// TIA Portal project "Lagerregal_3" (V20) (continued)
VERSION : 0.1
   VAR_INPUT
      eAutomatik : Bool;   // Automatikmodus
      eAusschalten : Bool;   // Ausschalten der Schrittkette
      T_1_2 : Bool;
      T_2_3 : Bool;
      T_3_4 : Bool := TRUE;
      T_4_5 : Bool := TRUE;
      T_5_6 : Bool := TRUE;
      T_6_7 : Bool := TRUE;
      T_7_8 : Bool := TRUE;
      T_8_9 : Bool := TRUE;
      T_9_10 : Bool := TRUE;
      T_10_1 : Bool := TRUE;
   END_VAR
   VAR_OUTPUT
      aSchrittnummer : Int;
   END_VAR
   VAR
      Step_1 : Bool;
      Step_2 : Bool;
      Step_3 : Bool;
      Step_4 : Bool;
      Step_5 : Bool;
      Step_6 : Bool;
      Step_7 : Bool;
      Step_8 : Bool;
      Step_9 : Bool;
      Step_10 : Bool;
   END_VAR
BEGIN

REGION Network 1: Step 1
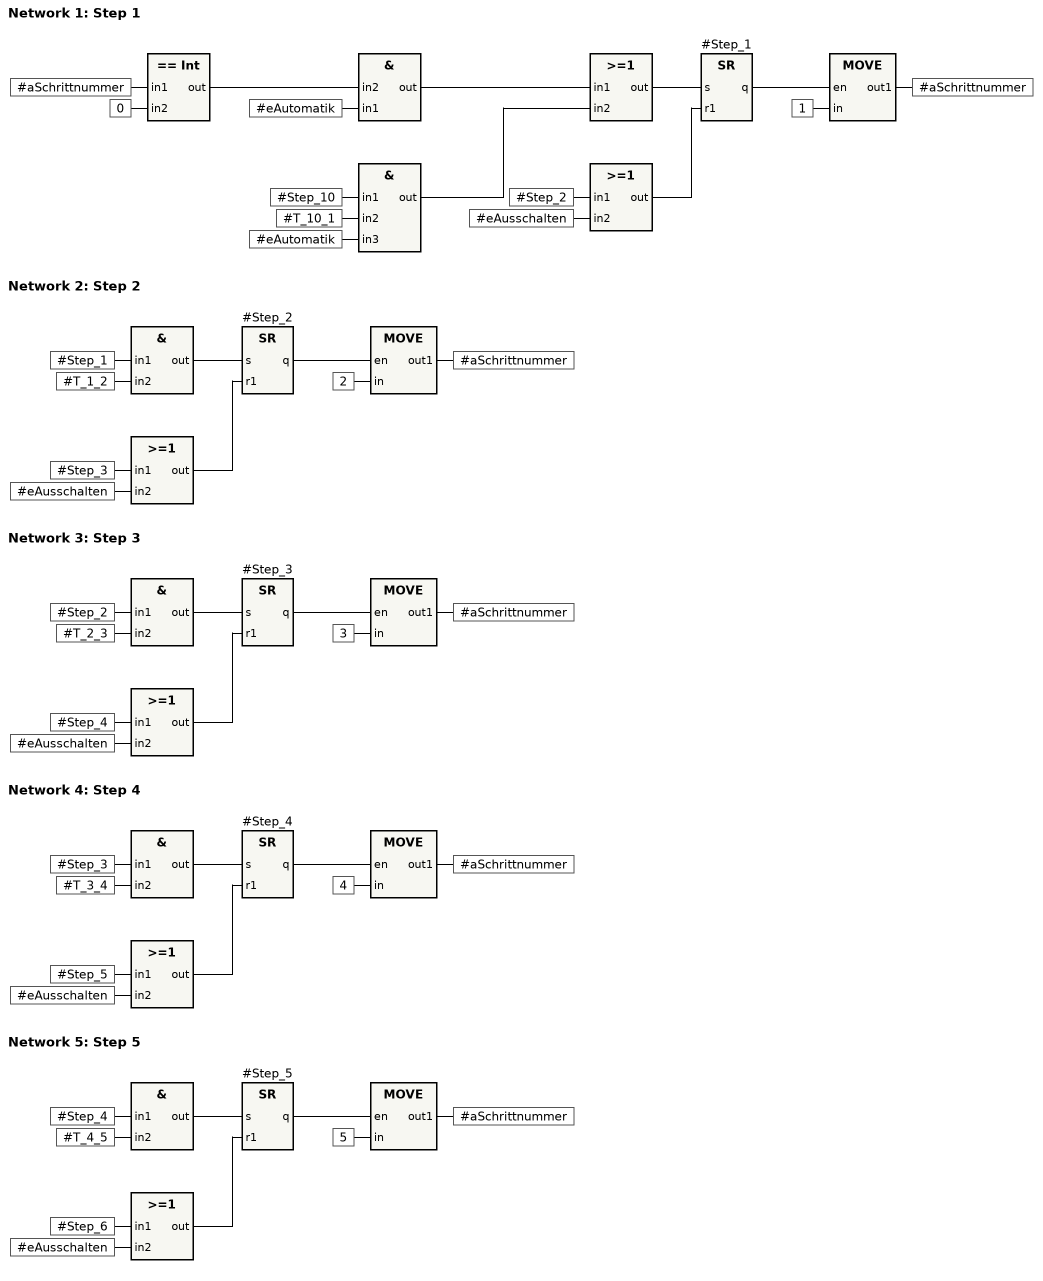
   IF ((#aSchrittnummer = 0) AND #eAutomatik) OR (#Step_10 AND #T_10_1 AND #eAutomatik) THEN
       #Step_1 := TRUE;   // SR flip-flop
   END_IF;
   IF #Step_2 OR #eAusschalten THEN #Step_1 := FALSE; END_IF;
   IF #Step_1 THEN #aSchrittnummer := 1; END_IF;
END_REGION

REGION Network 2: Step 2
   IF #Step_1 AND #T_1_2 THEN
       #Step_2 := TRUE;   // SR flip-flop
   END_IF;
   IF #Step_3 OR #eAusschalten THEN #Step_2 := FALSE; END_IF;
   IF #Step_2 THEN #aSchrittnummer := 2; END_IF;
END_REGION

REGION Network 3: Step 3
   IF #Step_2 AND #T_2_3 THEN
       #Step_3 := TRUE;   // SR flip-flop
   END_IF;
   IF #Step_4 OR #eAusschalten THEN #Step_3 := FALSE; END_IF;
   IF #Step_3 THEN #aSchrittnummer := 3; END_IF;
END_REGION

REGION Network 4: Step 4
   IF #Step_3 AND #T_3_4 THEN
       #Step_4 := TRUE;   // SR flip-flop
   END_IF;
   IF #Step_5 OR #eAusschalten THEN #Step_4 := FALSE; END_IF;
   IF #Step_4 THEN #aSchrittnummer := 4; END_IF;
END_REGION

REGION Network 5: Step 5
   IF #Step_4 AND #T_4_5 THEN
       #Step_5 := TRUE;   // SR flip-flop
   END_IF;
   IF #Step_6 OR #eAusschalten THEN #Step_5 := FALSE; END_IF;
   IF #Step_5 THEN #aSchrittnummer := 5; END_IF;
END_REGION

REGION Network 6: Step 6
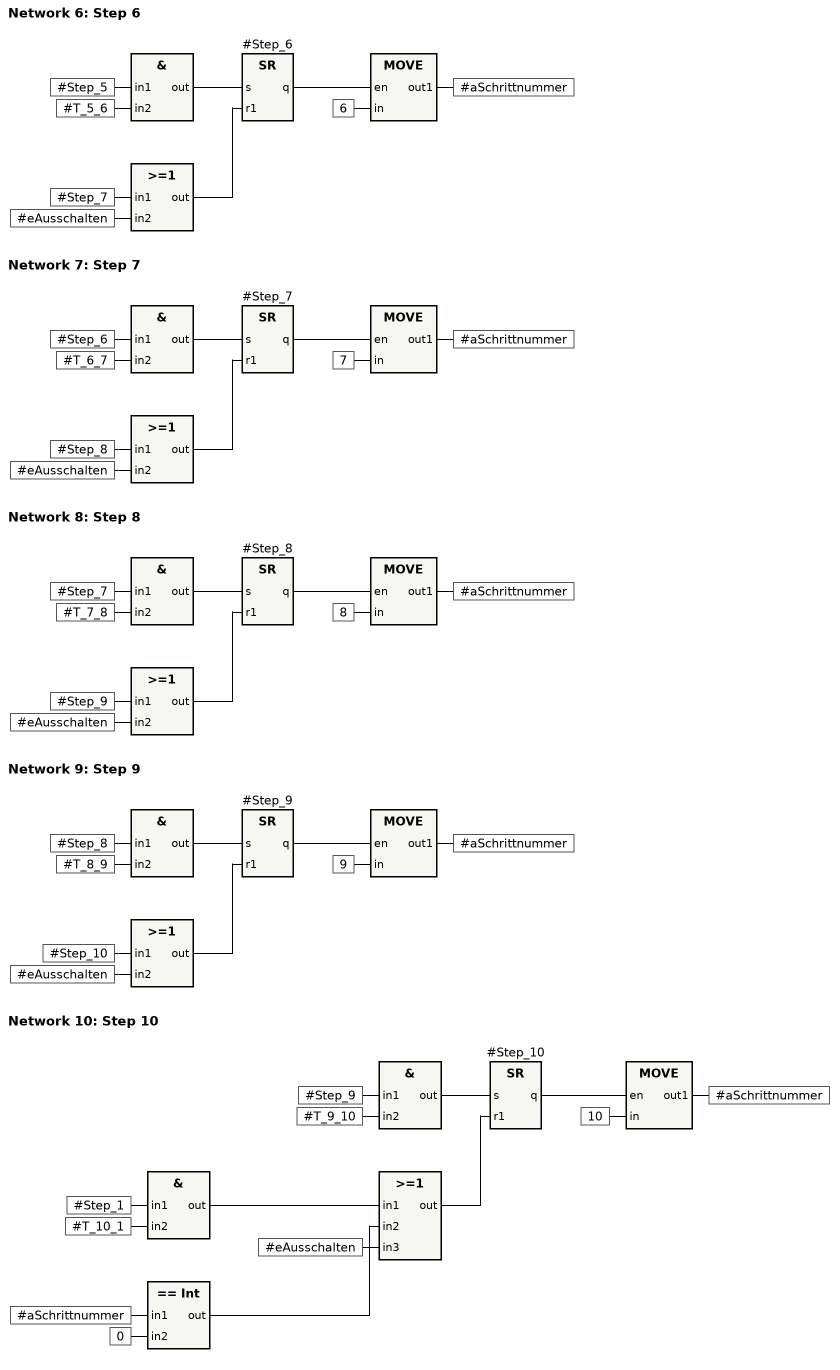
   IF #Step_5 AND #T_5_6 THEN
       #Step_6 := TRUE;   // SR flip-flop
   END_IF;
   IF #Step_7 OR #eAusschalten THEN #Step_6 := FALSE; END_IF;
   IF #Step_6 THEN #aSchrittnummer := 6; END_IF;
END_REGION

REGION Network 7: Step 7
   IF #Step_6 AND #T_6_7 THEN
       #Step_7 := TRUE;   // SR flip-flop
   END_IF;
   IF #Step_8 OR #eAusschalten THEN #Step_7 := FALSE; END_IF;
   IF #Step_7 THEN #aSchrittnummer := 7; END_IF;
END_REGION

REGION Network 8: Step 8
   IF #Step_7 AND #T_7_8 THEN
       #Step_8 := TRUE;   // SR flip-flop
   END_IF;
   IF #Step_9 OR #eAusschalten THEN #Step_8 := FALSE; END_IF;
   IF #Step_8 THEN #aSchrittnummer := 8; END_IF;
END_REGION

REGION Network 9: Step 9
   IF #Step_8 AND #T_8_9 THEN
       #Step_9 := TRUE;   // SR flip-flop
   END_IF;
   IF #Step_10 OR #eAusschalten THEN #Step_9 := FALSE; END_IF;
   IF #Step_9 THEN #aSchrittnummer := 9; END_IF;
END_REGION

REGION Network 10: Step 10
   IF #Step_9 AND #T_9_10 THEN
       #Step_10 := TRUE;   // SR flip-flop
   END_IF;
   IF (#Step_1 AND #T_10_1) OR (#aSchrittnummer = 0) OR #eAusschalten THEN #Step_10 := FALSE; END_IF;
   IF #Step_10 THEN #aSchrittnummer := 10; END_IF;
END_REGION

REGION Network 11: Schrittkette beenden, wenn der Automatikmodus beendet wird
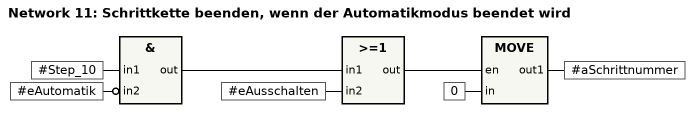
   IF (#Step_10 AND NOT #eAutomatik) OR #eAusschalten THEN #aSchrittnummer := 0; END_IF;
END_REGION
END_FUNCTION_BLOCK

FUNCTION "Aus_Anlage" : Void   // FC1, FBD
{ S7_Optimized_Access := 'TRUE' }
VERSION : 0.1
BEGIN

REGION Network 1 (SCL): Gabelsteuerung Kran_1
   "6M1" := "HMI_Schnittstelle".Ausgaenge."6M1";
   "6M2" := "HMI_Schnittstelle".Ausgaenge."6M2";
END_REGION

REGION Network 2 (SCL): Gabelsteuerung Kran_2
   "7M1" := "HMI_Schnittstelle".Ausgaenge."7M1";
   "7M2" := "HMI_Schnittstelle".Ausgaenge."7M2";
END_REGION

REGION Network 3 (SCL): Foerderbaender Einlass
   "1M1" := "HMI_Schnittstelle".Ausgaenge."1M1";
   "2M1" := "HMI_Schnittstelle".Ausgaenge."2M1";
   "3M1" := "HMI_Schnittstelle".Ausgaenge."3M1";
END_REGION

REGION Network 4 (SCL): Foerderbaender Auslass
   "4M1" := "HMI_Schnittstelle".Ausgaenge."4M1";
   "5M1" := "HMI_Schnittstelle".Ausgaenge."5M1";
END_REGION

REGION Network 5 (SCL): Leuchte Starttaster
   "HMI_Schnittstelle".Ausgaenge.H1 := "HMI_Schnittstelle".Eingaenge.S2;
END_REGION
END_FUNCTION

FUNCTION "Aus_HMI" : Void   // FC20, FBD
{ S7_Optimized_Access := 'TRUE' }
VERSION : 0.1
BEGIN
END_FUNCTION

FUNCTION "Aus_Kran" : Void   // FC30, SCL
{ S7_Optimized_Access := 'TRUE' }
VERSION : 0.1
   VAR_INPUT
      "eX-Soll" : Int;
      "eZ-Soll" : Int;
      eGabel_links : Bool;
      eGabel_rechts : Bool;
   END_VAR
   VAR_OUTPUT
      aKran_X : Int;
      aKran_Z : Int;
      aKran_Gabel_links : Bool;
      aKran_Gabel_rechts : Bool;
   END_VAR
BEGIN
   // Kran Gabel
   #aKran_Gabel_links := #eGabel_links;
   #aKran_Gabel_rechts := #eGabel_rechts;


   // Kran Position
   // Kran X-Soll-Position
   #"aKran_X" := #"eX-Soll";
   // Kran Z-Soll-Position
   #"aKran_Z" := #"eZ-Soll";
END_FUNCTION

FUNCTION "Ausgabe_Stapler_EIN" : Void   // FC70, FBD
{ S7_Optimized_Access := 'TRUE' }
VERSION : 0.1
BEGIN

REGION Network 1: Sollposition X
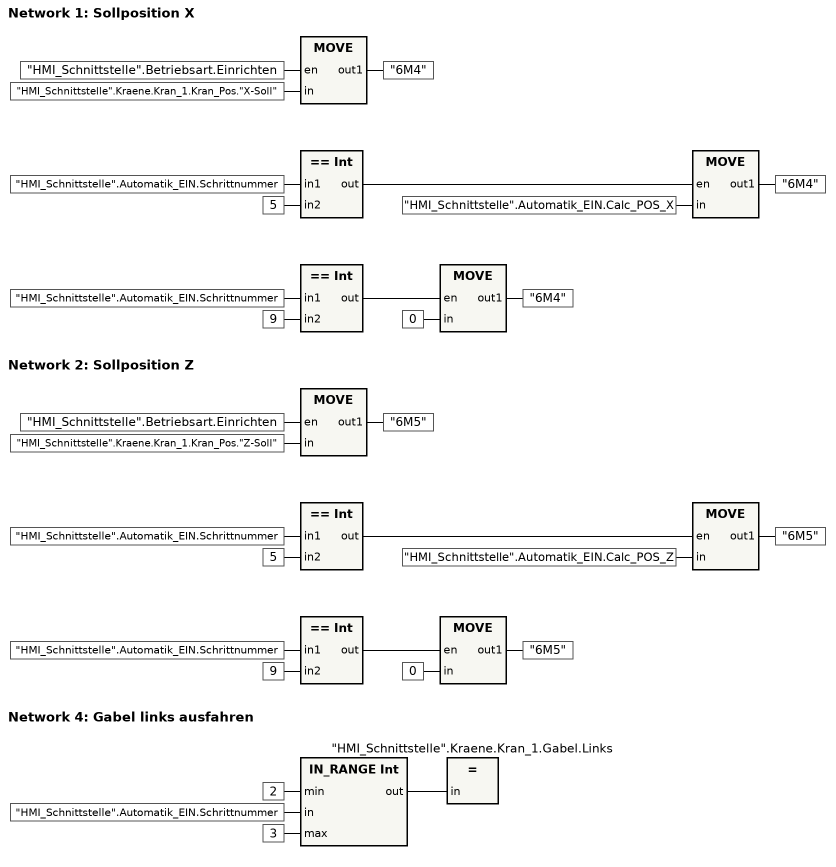
   IF "HMI_Schnittstelle".Betriebsart.Einrichten THEN
       "6M4" := "HMI_Schnittstelle".Kraene.Kran_1.Kran_Pos."X-Soll";
   END_IF;
   IF "HMI_Schnittstelle".Automatik_EIN.Schrittnummer = 5 THEN
       "6M4" := "HMI_Schnittstelle".Automatik_EIN.Calc_POS_X;
   END_IF;
   IF "HMI_Schnittstelle".Automatik_EIN.Schrittnummer = 9 THEN "6M4" := 0; END_IF;
END_REGION

REGION Network 2: Sollposition Z
   IF "HMI_Schnittstelle".Betriebsart.Einrichten THEN
       "6M5" := "HMI_Schnittstelle".Kraene.Kran_1.Kran_Pos."Z-Soll";
   END_IF;
   IF "HMI_Schnittstelle".Automatik_EIN.Schrittnummer = 5 THEN
       "6M5" := "HMI_Schnittstelle".Automatik_EIN.Calc_POS_Z;
   END_IF;
   IF "HMI_Schnittstelle".Automatik_EIN.Schrittnummer = 9 THEN "6M5" := 0; END_IF;
END_REGION

REGION Network 3 (SCL): Z-Achse Kran 1 Soll-Pos
   // Einrichtbetrieb
   IF "HMI_Schnittstelle".Betriebsart.Einrichten THEN
       "6M5" := "HMI_Schnittstelle".Kraene.Kran_1.Kran_Pos."Z-Soll";

   // Automatikbetrieb    
   ELSIF "HMI_Schnittstelle".Automatik_EIN.Schrittnummer = 3 THEN
       // Palette aus Grundstellung anheben
       "6M5" := "Anheben_Absenken" + 2;
   ELSIF "HMI_Schnittstelle".Automatik_EIN.Schrittnummer = 5 THEN
       //Fach mit Nummer anfahren
       "6M5" := "HMI_Schnittstelle".Automatik_EIN.Calc_POS_Z;
   ELSIF "HMI_Schnittstelle".Automatik_EIN.Schrittnummer = 7 THEN
       // Palette in Regal einlagern
       "6M5" := "HMI_Schnittstelle".Automatik_EIN.Calc_POS_Z - "Anheben_Absenken";
   ELSIF "HMI_Schnittstelle".Automatik_EIN.Schrittnummer = 9 THEN
       // Stapler in Grundstellung
       "6M5" := 0;
   END_IF;
END_REGION

REGION Network 4: Gabel links ausfahren
   "HMI_Schnittstelle".Kraene.Kran_1.Gabel.Links := (2 <= "HMI_Schnittstelle".Automatik_EIN.Schrittnummer) AND ("HMI_Schnittstelle".Automatik_EIN.Schrittnummer <= 3);
END_REGION

REGION Network 5 (SCL): Gabel rechts ausfahren
   "HMI_Schnittstelle".Kraene.Kran_1.Gabel.Rechts := "HMI_Schnittstelle".Automatik_EIN.Schrittnummer = 6
                                                   OR "HMI_Schnittstelle".Automatik_EIN.Schrittnummer = 7;
END_REGION
END_FUNCTION

FUNCTION "Berechne_Offset" : Void   // FC5000, SCL
{ S7_Optimized_Access := 'TRUE' }
VERSION : 0.1
   VAR_INPUT
      eFach_Nr : DInt;
      eFach_Anzahl : DInt;
      eFach_Breite : DInt;
      eFach_Hoehe : DInt;
      eOffset_X : DInt;
      eOffset_Z : DInt;
   END_VAR
   VAR_OUTPUT
      aPos_X : DInt;
      aPos_Z : DInt;
   END_VAR
BEGIN
   (*
      Der Baustein berechnet die Koordinaten (X,Z) eines Fachs
      in Abhängigkeit von einer Fachnummer

      Der Baustein ist universell einsetzbar für alle gleichhbleibenden Raster.
   *)

   // Position setzen
   IF #eFach_Nr > 0 THEN
       #aPos_X := ((#eFach_Nr - 1) MOD #eFach_Anzahl) * #eFach_Breite + #eOffset_X;
       #aPos_Z := ((#eFach_Nr - 1) / #eFach_Anzahl) * #eFach_Hoehe + #eOffset_Z;
   ELSE
       #aPos_X := #aPos_Z := 0;
   END_IF;
END_FUNCTION

ORGANIZATION_BLOCK "Main"   // OB1, FBD, ProgramCycle
TITLE = "Main Program Sweep (Cycle)"
{ S7_Optimized_Access := 'TRUE' }
VERSION : 0.1
   VAR_INPUT
      Initial_Call : Bool;   // Initial call of this OB
      Remanence : Bool;   // =True, if remanent data are available
   END_VAR
BEGIN

REGION Network 1: Anlage
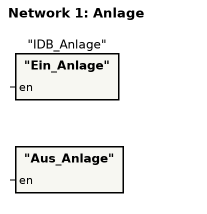
   "IDB_Anlage"();   // "Ein_Anlage"
   "Aus_Anlage"();
END_REGION
END_ORGANIZATION_BLOCK

ORGANIZATION_BLOCK "Main_einlagern"   // OB123, FBD, ProgramCycle
TITLE = "Main Program Sweep (Cycle)"
{ S7_Optimized_Access := 'TRUE' }
VERSION : 0.1
   VAR_INPUT
      Initial_Call : Bool;   // Initial call of this OB
      Remanence : Bool;   // =True, if remanent data are available
   END_VAR
BEGIN

REGION Network 1: Test ob Kran in Grundstellung ist
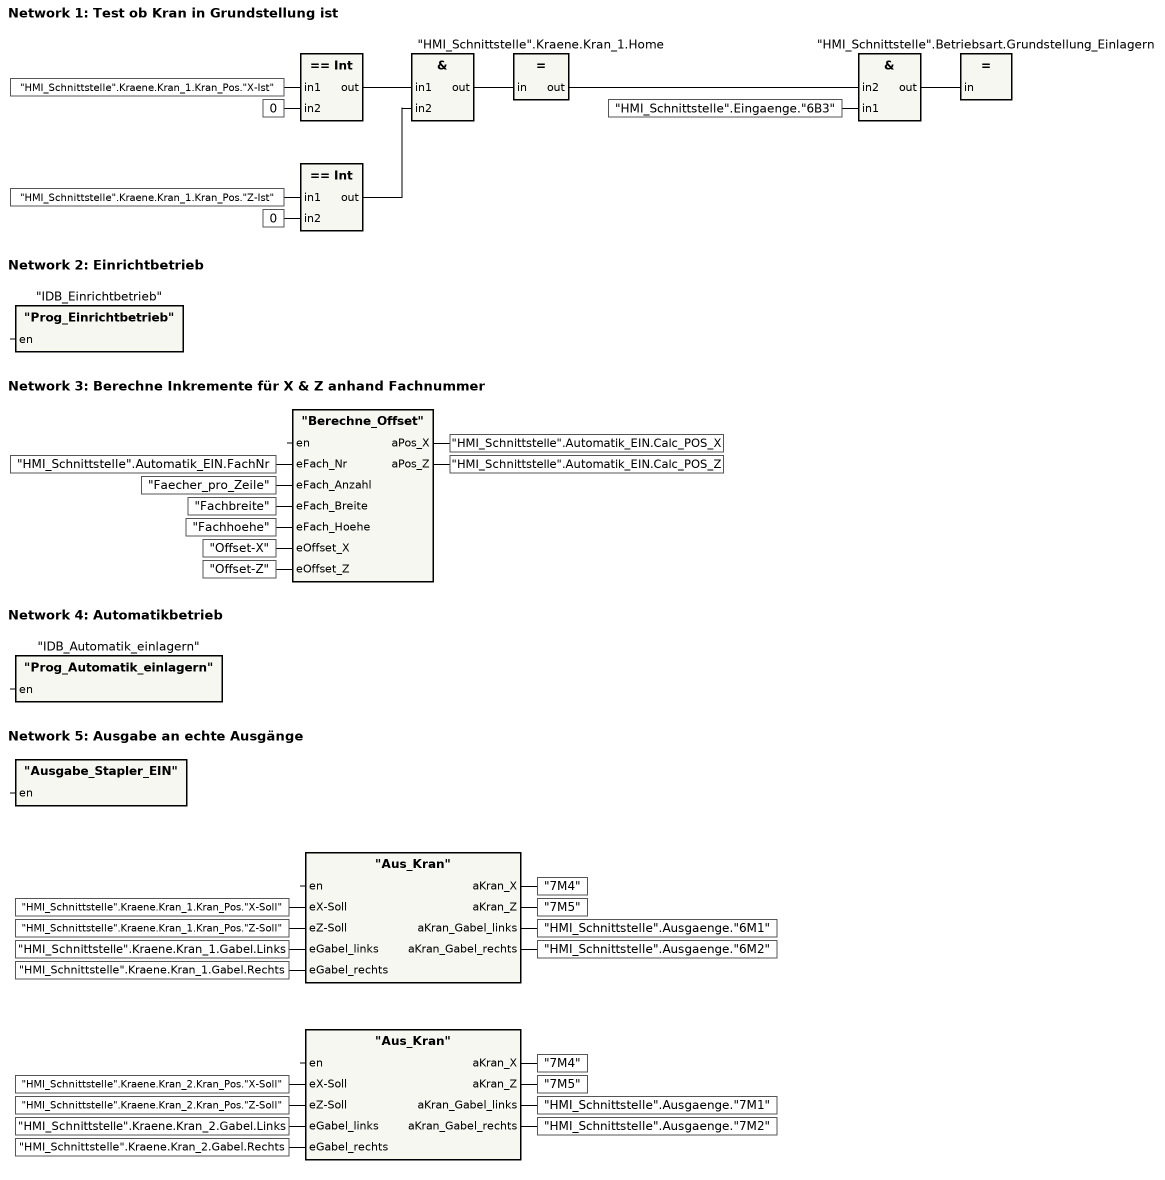
   "HMI_Schnittstelle".Kraene.Kran_1.Home := ("HMI_Schnittstelle".Kraene.Kran_1.Kran_Pos."X-Ist" = 0) AND ("HMI_Schnittstelle".Kraene.Kran_1.Kran_Pos."Z-Ist" = 0);
   "HMI_Schnittstelle".Betriebsart.Grundstellung_Einlagern := "HMI_Schnittstelle".Kraene.Kran_1.Home AND "HMI_Schnittstelle".Eingaenge."6B3";
END_REGION

REGION Network 2: Einrichtbetrieb
   "IDB_Einrichtbetrieb"();   // "Prog_Einrichtbetrieb"
END_REGION

REGION Network 3: Berechne Inkremente für X & Z anhand Fachnummer
   "Berechne_Offset"(eFach_Nr := "HMI_Schnittstelle".Automatik_EIN.FachNr,
                     eFach_Anzahl := "Faecher_pro_Zeile",
                     eFach_Breite := "Fachbreite",
                     eFach_Hoehe := "Fachhoehe",
                     eOffset_X := "Offset-X",
                     eOffset_Z := "Offset-Z",
                     aPos_X => "HMI_Schnittstelle".Automatik_EIN.Calc_POS_X,
                     aPos_Z => "HMI_Schnittstelle".Automatik_EIN.Calc_POS_Z);
END_REGION

REGION Network 4: Automatikbetrieb
   "IDB_Automatik_einlagern"();   // "Prog_Automatik_einlagern"
END_REGION

REGION Network 5: Ausgabe an echte Ausgänge
   "Ausgabe_Stapler_EIN"();
   "Aus_Kran"("eX-Soll" := "HMI_Schnittstelle".Kraene.Kran_1.Kran_Pos."X-Soll",
              "eZ-Soll" := "HMI_Schnittstelle".Kraene.Kran_1.Kran_Pos."Z-Soll",
              eGabel_links := "HMI_Schnittstelle".Kraene.Kran_1.Gabel.Links,
              eGabel_rechts := "HMI_Schnittstelle".Kraene.Kran_1.Gabel.Rechts,
              aKran_X => "7M4",
              aKran_Z => "7M5",
              aKran_Gabel_links => "HMI_Schnittstelle".Ausgaenge."6M1",
              aKran_Gabel_rechts => "HMI_Schnittstelle".Ausgaenge."6M2");
   "Aus_Kran"("eX-Soll" := "HMI_Schnittstelle".Kraene.Kran_2.Kran_Pos."X-Soll",
              "eZ-Soll" := "HMI_Schnittstelle".Kraene.Kran_2.Kran_Pos."Z-Soll",
              eGabel_links := "HMI_Schnittstelle".Kraene.Kran_2.Gabel.Links,
              eGabel_rechts := "HMI_Schnittstelle".Kraene.Kran_2.Gabel.Rechts,
              aKran_X => "7M4",
              aKran_Z => "7M5",
              aKran_Gabel_links => "HMI_Schnittstelle".Ausgaenge."7M1",
              aKran_Gabel_rechts => "HMI_Schnittstelle".Ausgaenge."7M2");
END_REGION

REGION Network 6: Test ob Kran in Bewegung ist
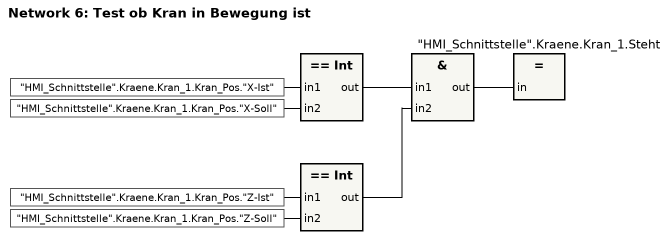
   "HMI_Schnittstelle".Kraene.Kran_1.Steht := ("HMI_Schnittstelle".Kraene.Kran_1.Kran_Pos."X-Ist" = "HMI_Schnittstelle".Kraene.Kran_1.Kran_Pos."X-Soll") AND ("HMI_Schnittstelle".Kraene.Kran_1.Kran_Pos."Z-Ist" = "HMI_Schnittstelle".Kraene.Kran_1.Kran_Pos."Z-Soll");
END_REGION
END_ORGANIZATION_BLOCK

(* ===== HMI "HMI_RT_1" =====
system functions are stored by id; their names below are inferred from use
connection "HMI_Verbindung_1": ETHERNET, S7_1500_OMS

HMI tags "Standard-Variablentabelle"
   "HMI_Schnittstelle_Kraene_Kran_1_Z-Soll" : Int = PLC HMI_Schnittstelle.Kraene.Kran_1.Kran_Pos.Z-Soll, 1 s
   "HMI_Schnittstelle_Kraene_Kran_1_X-Soll" : Int = PLC HMI_Schnittstelle.Kraene.Kran_1.Kran_Pos.X-Soll, 1 s
   "HMI_Schnittstelle_Kraene_Kran_1_X-Ist" : Int = PLC HMI_Schnittstelle.Kraene.Kran_1.Kran_Pos.X-Ist, 1 s
   "HMI_Schnittstelle_Kraene_Kran_1_Z-Ist" : Int = PLC HMI_Schnittstelle.Kraene.Kran_1.Kran_Pos.Z-Ist, 1 s
   "HMI_Schnittstelle_HMI_X-Neg" : Bool = PLC HMI_Schnittstelle.HMI.X-Neg, 1 s
   "HMI_Schnittstelle_HMI_X-Pos" : Bool = PLC HMI_Schnittstelle.HMI.X-Pos, 1 s
   "HMI_Schnittstelle_HMI_Z-Neg" : Bool = PLC HMI_Schnittstelle.HMI.Z-Neg, 1 s
   "HMI_Schnittstelle_HMI_Z-Pos" : Bool = PLC HMI_Schnittstelle.HMI.Z-Pos, 1 s
   "HMI_Schnittstelle_HMI_Inkrement" : UInt = PLC HMI_Schnittstelle.HMI.Inkrement, 1 s
   "HMI_Schnittstelle_Ausgaenge_Fach_ansteuern" : Bool = PLC HMI_Schnittstelle.Fach_ansteuern, 1 s
   "HMI_Schnittstelle_Ausgaenge_Fach" : Int = PLC HMI_Schnittstelle.Fach, 1 s
   "Clock_1Hz" : Bool = PLC Clock_1Hz AT %M0.5, 100 ms
   "HMI_Schnittstelle_Fach" : Int = PLC HMI_Schnittstelle.Fach, 1 s
   "HMI_Schnittstelle_Fach_ansteuern" : Bool = PLC HMI_Schnittstelle.Fach_ansteuern, 1 s
   "Warenlager_Lager{1}_Flags_Belegt" : Bool = PLC Warenlager.Lager[1].Flags.Belegt, 1 s
   "Warenlager_Lager{1}_Flags_In_Benutzung" : Bool = PLC Warenlager.Lager[1].Flags.In_Benutzung, 1 s

screen "Lageransicht" 800x420, template "Menüleiste"
   Button "Schaltfläche_4" at 10,438 size 96x32; TextOff 'Teachen'
      on Press: ActivateScreen("Teachmodus", 0)
   Rectangle "Rechteck_1" at 650,280 size 50x50
      Appearance <- "Warenlager_Lager{1}_Flags_Belegt"
   TextField "Textfeld_1" at 650,280 size 50x50; Text '1'
      Appearance <- "Warenlager_Lager{1}_Flags_In_Benutzung"

screen "Teachmodus" 800x420, template "Menüleiste"
   Button "Schaltfläche_1" at 694,10 size 96x32; TextOff 'Zurück'
      on Press: function_efd93a16()
   TextField "Textfeld_1" at 308,10 size 184x23; Text 'Kalibrierungsmodus'
   Slider "Schieberegler_2" at 113,300 size 230x50; Caption 'Breite'
      ProcessValue <- "HMI_Schnittstelle_Kraene_Kran_1_X-Soll"
   IOField "EA-Feld_8" at 370,67 size 96x32; FormatPattern 99999
      ProcessValue <- "HMI_Schnittstelle_Kraene_Kran_1_X-Ist"
   IOField "EA-Feld_9" at 485,68 size 96x32; FormatPattern 99999
      ProcessValue <- "HMI_Schnittstelle_Kraene_Kran_1_Z-Ist"
   Slider "Schieberegler_1" at 10,37 size 50x230; Caption 'Höhe'
      ProcessValue <- "HMI_Schnittstelle_Kraene_Kran_1_Z-Soll"
   Button "Schaltfläche_5" at 345,300 size 25x50; TextOff '-'
      on Press: function_b14e0dd5("HMI_Schnittstelle_HMI_X-Neg", 0)
      Appearance <- "HMI_Schnittstelle_HMI_X-Neg"
   IOField "EA-Feld_7" at 10,300 size 70x50; FormatPattern 99999
      ProcessValue <- "HMI_Schnittstelle_HMI_Inkrement"
   Button "Schaltfläche_7" at 10,269 size 50x25; TextOff '-'
      on Press: function_b14e0dd5("HMI_Schnittstelle_HMI_Z-Neg", 0)
      Appearance <- "HMI_Schnittstelle_HMI_Z-Neg"
   Button "Schaltfläche_8" at 10,10 size 50x25; TextOff '+'
      on Press: function_b14e0dd5("HMI_Schnittstelle_HMI_Z-Pos", 0)
      Appearance <- "HMI_Schnittstelle_HMI_Z-Pos"
   Button "Schaltfläche_6" at 86,300 size 25x50; TextOff '+'
      on Press: function_b14e0dd5("HMI_Schnittstelle_HMI_X-Pos", 0)
      Appearance <- "HMI_Schnittstelle_HMI_X-Pos"
   TextField "Textfeld_2" at 370,42 size 111x23; Text 'Ist-X-Achse'
   TextField "Textfeld_3" at 485,42 size 110x23; Text 'Ist-Z-Achse'
   TextField "Textfeld_4" at 370,103 size 88x23; Text 'Fach-Nr.:'
   IOField "EA-Feld_1" at 370,128 size 96x32; FormatPattern 99
      ProcessValue <- "HMI_Schnittstelle_Fach"
   Button "Schaltfläche_2" at 485,128 size 96x32; TextOff 'Testen'
      on Press: function_b14e0dd5("HMI_Schnittstelle_Fach_ansteuern", 0)

screen "Detailansicht" 800x420, template "Menüleiste"
   Button "Schaltfläche_1" at 694,10 size 96x32; TextOff 'Zurück'
      on Press: function_efd93a16()

Template "Menüleiste" 800x420
   Button "Vorlage_Schaltfläche_1" at 0,360 size 80x60; TextOff 'HOME'
      on Click: ActivateScreen("Lageransicht", 0)
   Button "Vorlage_Schaltfläche_2" at 80,360 size 80x60; TextOff 'Text'
      on Click: ActivateScreen("Lageransicht", 0)
   Button "Vorlage_Schaltfläche_3" at 160,360 size 80x60; TextOff 'Text'
      on Click: ActivateScreen("Lageransicht", 0)
   Button "Vorlage_Schaltfläche_4" at 240,360 size 80x60; TextOff 'Text'
      on Click: ActivateScreen("Lageransicht", 0)
   Button "Vorlage_Schaltfläche_5" at 320,360 size 80x60; TextOff 'TEACH'
      on Click: ActivateScreen("Teachmodus", 0)
   Button "Vorlage_Schaltfläche_6" at 400,360 size 80x60; TextOff 'Text'
      on Click: ActivateScreen("Lageransicht", 0)
   Button "Vorlage_Schaltfläche_7" at 480,360 size 80x60; TextOff 'Text'
      on Click: ActivateScreen("Lageransicht", 0)
   Button "Vorlage_Schaltfläche_8" at 560,360 size 80x60; TextOff 'Text'
      on Click: ActivateScreen("Lageransicht", 0)
   Button "Vorlage_Schaltfläche_9" at 640,360 size 80x60; TextOff 'Text'
      on Click: ActivateScreen("Lageransicht", 0)
   Button "Vorlage_Schaltfläche_10" at 720,360 size 80x60; TextOff 'Text'
      on Click: ActivateScreen("Lageransicht", 0)
*)